// TIA Portal project "e009004v441" (V15.1)

(* hardware
DEVICE "Roll Forming"  TP1200 Comfort
   slot 0: "Roll Forming"  TP1200 Comfort  6AV2 124-0MC01-0AX0  15.1.0.0
   slot 1: "HMI_RT_1"  TP1200 Comfort  6AV2 124-0MC01-0AX0  15.1.0.0
   slot 5: "Roll Forming.IE_CP_1"  PROFINET Interface  15.0.1.0
      slot 1: "Interfaz PROFINET_1"  PROFINET Interface
         slot 1: "Port_1"  Port
         slot 2: "Port_2"  Port
   slot 7: "Roll Forming.MPI/DP_CP_1"  MPI/DP Interface  15.0.1.0
DEVICE "Dispositivo GSD_1"  GSD.Device
   slot 0: "Rack_0"  Rail
   slot 0: "Perfiladora"  6SL3 040-1MA00-0xxx  V4.3
DEVICE "PC-System_1"  SIMATIC PC station
   slot 0: "Estación PC SIMATIC"  Rail  SIMATIC PC-Station  V1.0
      slot 125: "Stationmanager"  Station_Manager  V6.0.4
   slot 1: "HMI_RT_2"  WinCC RT Advanced  6AV2 104-0xxxx-xxxx  15.1.0.0
      slot 33792: "Interfaz host"  Host interface
*)

(* ===== HMI "HMI_RT_1" =====

ScreenModuleEditorView "Bloc affichage_2" 800x600
   GraphicView "Affichage graphique" at 10,10 size 40x80; Picture "Graphique_9"
*)

(* ===== HMI "HMI_RT_1" =====
system functions are stored by id; their names below are inferred from use
connection "CPU 313C-2 DP": IF1 B, SIMATIC S7 300/400 MPI

HMI tags "Tabla de variables estándar"
   "DB_OP.COD2_ARRET" : DInt AT %DB50.DBD138, 1 s   // Encoder Formador 2 : Parar 1/10 mm
   "Desactivar_Falla59" : Bool AT %M87.2, 1 s
   "Desactivar_Falla78" : Bool AT %M89.5, 1 s
   "Desactivar_Falla47" : Bool AT %M85.6, 1 s
   "Desactivar_Falla84" : Bool AT %M90.3, 1 s
   "DB_OP.ACQ_DEFAUT" : Bool AT %DB50.DBX0.1, 1 s
   "Desactivar_Falla58" : Bool AT %M87.1, 1 s
   "Desactivar_Falla75" : Bool AT %M89.2, 1 s
   "35S2" : Bool AT %I12.1, 1 s   // Plegador 2 Fijación Abajo
   "28S3" : Bool AT %I5.2, 1 s   // Formador Herramienta 2 Matriz Off
   "Desactivar_Falla104" : Bool AT %M92.7, 1 s
   "Desactivar_Falla3" : Bool AT %M80.2, 1 s
   "Alarma_Cinta" : Bool AT %M96.4, 1 s
   "Desactivar_Falla68" : Bool AT %M88.3, 1 s
   "Desactivar_Falla38" : Bool AT %M84.5, 1 s
   "28S2" : Bool AT %I5.1, 1 s   // Formador Herramienta 2 Martillo On
   "DB_OP.COD1_VAL" : DInt AT %DB50.DBD100, 1 s   // Encoder Perfilador 1 : Valor 1/10 mm
   "31S3" : Bool AT %I8.2, 1 s   // Descargador Atrás
   "25S4" : Bool AT %I2.3, 1 s   // Pistón 1 Araña Contraído
   "Desactivar_Falla80" : Bool AT %M89.7, 1 s
   "Desactivar_Falla119" : Bool AT %M94.6, 1 s
   "Desactivar_Falla88" : Bool AT %M90.7, 1 s
   "HeladerasxMin" : Real AT %MD132, 1 s
   "Desactivar_Falla52" : Bool AT %M86.3, 1 s
   "Alarma_General" : Bool AT %M97.1, 1 s
   "DB_OP.DB_VAR" : Array [0..20] of Int AT %DB50.DBX8.0, 1 s   // Variables temporales
   "Desactivar_Falla11" : Bool AT %M81.2, 1 s
   "DB_OP.PI_COD_VAL" : DInt AT %DB50.DBD300, 1 s   // Encóder Pinza : Valor 1/10 mm
   "Desactivar_Falla116" : Bool AT %M94.3, 1 s
   "Desactivar_Falla102" : Bool AT %M92.5, 1 s
   "Hab_Medición" : Bool AT %M102.6, 1 s
   "35S3b" : Bool AT %I15.6, 1 s   // Plegador 2 posición Arriba (pata)
   "DB_OP.COD1_INIT" : DInt AT %DB50.DBD116, 1 s   // Encoder Perfilador 1 : Consigna Inicial 1/10 mm
   "Desactivar_Falla92" : Bool AT %M91.3, 1 s
   "28S8" : Bool AT %I5.7, 1 s   // Ajuste Formador Fin de Carrera Máx.
   "31S7b" : Bool AT %I15.5, 1 s   // Plegador 1 posición Arriba (pata)
   "DB_OP.COD2_CONS" : DInt AT %DB50.DBD134, 1 s   // Encoder Formador 2 : Consigna Posición 1/10 mm
   "DB_OP.DEF08" : Int AT %DB50.DBW94, 1 s   // IMAGE DEFAUT DBW 64
   "23S4" : Bool AT %I0.7, 1 s   // Presostato Freno Perfilador
   "Desactivar_Falla25" : Bool AT %M83.0, 1 s
   "Desactivar_Falla56" : Bool AT %M86.7, 1 s
   "DB_OP.DF_QM01" : Bool AT %DB50.DBX50.2, 1 s   // Térmico Intercambiador de Chapas
   "DB_OP.DEF06" : Int AT %DB50.DBW90, 1 s   // IMAGE DEFAUT DBW 60
   "DI8_CU_PL" : Bool AT %I62.7, 1 s   // Entrada Digital 8 CU Plegadores
   "DB_OP.DF_QM14" : Bool AT %DB50.DBX50.1, 1 s   // Térmico Calentador de Chapa
   "Desactivar_Falla39" : Bool AT %M84.6, 1 s
   "DB_OP.DEF01" : Int AT %DB50.DBW80, 1 s   // IMAGE DEFAUT DBW 50
   "32S5" : Bool AT %I9.4, 1 s   // Plegador 1 Extensión 2 Prensa Abajo
   "35S4_0" : Bool AT %I12.3, 1 s   // Plegador 2 Abajo
   "Desactivar_Falla112" : Bool AT %M93.7, 1 s
   "29S5" : Bool AT %I6.4, 1 s   // Pinza Cerrada
   "25S3" : Bool AT %I2.2, 1 s   // Fin de Carrera Araña Arriba
   "Desactivar_Falla93" : Bool AT %M91.4, 1 s
   "Desactivar_Falla111" : Bool AT %M93.6, 1 s
   "DB_OP.DF_QM06" : Bool AT %DB50.DBX51.2, 1 s   // Térmico Grupo Hidráulico Freno Perfilador
   "DB_OP.DF_VAR02" : Bool AT %DB50.DBX50.3, 1 s   // Defecto Vaiador Araña
   "30S3" : Bool AT %I7.2, 1 s   // Plegadora Tenaza arriba
   "Desactivar_Falla10" : Bool AT %M81.1, 1 s
   "DB_OP.PL2_COD_COEF" : Real AT %DB50.DBD262, 1 s   // Encoder Plegador 2 : Coeficiente Corrección
   "Desactivar_Falla6" : Bool AT %M80.5, 1 s
   "35S3" : Bool AT %I12.2, 1 s   // Plegador 2 Arriba
   "Desactivar_Falla103" : Bool AT %M92.6, 1 s
   "Alarma_Plegador" : Bool AT %M96.7, 1 s
   "DB_OP.PI_COD_DEC_PLI" : DInt AT %DB50.DBD322, 1 s   // Encóder Pinza : DECALAGE OUTIL PLIEUSE 1/10 mm
   "Desactivar_Falla36" : Bool AT %M84.3, 1 s
   "DB_OP.DF_LIM_PL1" : Bool AT %DB50.DBX51.7, 1 s   // Defecto Límite Plegador 1
   "Desactivar_Falla16" : Bool AT %M81.7, 1 s
   "26S4" : Bool AT %I3.3, 1 s   // Bajar Velocidad Transporte de Araña para Tomar Chapa
   "35S7" : Bool AT %I12.6, 1 s   // Plegador 2 Extensión 1 Prensa Abajo
   "27S4" : Bool AT %I4.3, 1 s   // Chapa en salida Perfilador
   "DB_OP.P_DEFAUT" : Bool AT %DB50.DBX0.0, 1 s
   "Desactivar_Falla71" : Bool AT %M88.6, 1 s
   "Desactivar_Falla48" : Bool AT %M85.7, 1 s
   "Desactivar_Falla125" : Bool AT %M95.4, 1 s
   "26S1" : Bool AT %I3.0, 1 s   // Tulipas no apoyadas en Chapa
   "DB_OP.COD1_CMD" : Bool AT %DB50.DBX128.0, 1 s   // Encoder Perfilador 1 : Inicio
   "30S7" : Bool AT %I7.6, 1 s   // Plegador 1 Cepillos Arriba
   "Desactivar_Falla83" : Bool AT %M90.2, 1 s
   "Alarma_Formador" : Bool AT %M96.5, 1 s
   "DB_OP.DEF05" : Int AT %DB50.DBW88, 1 s   // IMAGE DEFAUT DBW 58
   "Desactivar_Falla100" : Bool AT %M92.3, 1 s
   "21S6" : Bool AT %I124.7, 1 s   // Alineador Eje X Plegador 1 OFF
   "47K4" : Bool AT %Q8.3, 1 s   // Plegador 2 Bajar
   "Tiempo_Heladera_Prom" : Real AT %DB1.DBD40, 1 s
   "Desactivar_Falla107" : Bool AT %M93.2, 1 s
   "Desactivar_Falla114" : Bool AT %M94.1, 1 s
   "Desactivar_Falla21" : Bool AT %M82.4, 1 s
   "Desactivar_Falla31" : Bool AT %M83.6, 1 s
   "36S5" : Bool AT %I13.6, 1 s   // Plegador 2 Cepillos Arriba
   "29S4" : Bool AT %I6.3, 1 s   // Pinza Abierta
   "Desactivar_Falla97" : Bool AT %M92.0, 1 s
   "Desactivar_Falla14" : Bool AT %M81.5, 1 s
   "Desactivar_Falla82" : Bool AT %M90.1, 1 s
   "DB_OP.DF_LIM_PL2" : Bool AT %DB50.DBX52.0, 1 s   // Defecto Límite Plegador 2
   "Desactivar_Falla110" : Bool AT %M93.5, 1 s
   "35S2_0" : Bool AT %I12.1, 1 s   // Plegador 2 Fijación Abajo
   "Desactivar_Falla109" : Bool AT %M93.4, 1 s
   "Desactivar_Falla95" : Bool AT %M91.6, 1 s
   "36S6" : Bool AT %I13.7, 1 s   // Plegador 2 Cepillos Abajo
   "Desactivar_Falla76" : Bool AT %M89.3, 1 s
   "Selec_Pleg" : Int, internal
   "31S8" : Bool AT %I8.7, 1 s   // Plegador 1 Abajo
   "Alarma_Rolos" : Bool AT %M96.2, 1 s
   "27S6" : Bool AT %I4.5, 1 s   // Formador Herramienta 1 Martillo On
   "30S2" : Bool AT %I7.1, 1 s   // Plegadora Tenaza atrás
   "30S1" : Bool AT %I7.0, 1 s   // Plegadora Tenaza adelante
   "25S5" : Bool AT %I2.4, 1 s   // Fin de Carrera Araña Abajo
   "Desactivar_Falla29" : Bool AT %M83.4, 1 s
   "Desactivar_Falla13" : Bool AT %M81.4, 1 s
   "Desactivar_Falla23" : Bool AT %M82.6, 1 s
   "Alarma_Descargador" : Bool AT %M97.0, 1 s
   "DB_OP.PL1_COD_OFFSET" : DInt AT %DB50.DBD208, 1 s   // Encoder Plegador 1 : Consigna Inicial 1/10 mm
   "30S8" : Bool AT %I7.7, 1 s   // Plegador 1 Cepillos Abajo
   "DB_OP.PL2_COD_OFFSET" : DInt AT %DB50.DBD258, 1 s   // Encoder Plegador 2 : Consigna Inicial 1/10 mm
   "DB_OP.PI_COD_DEC_FORM" : DInt AT %DB50.DBD318, 1 s   // Encóder Pinza : DECALAGE OUTIL FORMAGE 1/10 mm
   "Alarma_Araña" : Bool AT %M96.1, 1 s
   "oHomming" : Bool AT %Q9.2, 1 s   // Lámpara Homming realizado
   "26S7" : Bool AT %I3.6, 1 s   // Presencia de Almacén 2 en Puesto de Trabajo
   "Simu Suelta Chapa" : Bool AT %M65.1, 1 s
   "Desactivar_Falla108" : Bool AT %M93.3, 1 s
   "DB_OP.COD2_COEF" : Real AT %DB50.DBD150, 1 s   // Encoder Formador 2 : Coeficiente Corrección
   "Ver_Tendencia" : Bool, internal
   "Desactivar_Falla46" : Bool AT %M85.5, 1 s
   "Desactivar_Falla40" : Bool AT %M84.7, 1 s
   "Simu Toma Chapa" : Bool AT %M65.0, 1 s
   "32S6" : Bool AT %I9.5, 1 s   // Plegador 1 Extensión 2 Prensa Arriba
   "Desactivar_Falla69" : Bool AT %M88.4, 1 s
   "35S3_0" : Bool AT %I12.2, 1 s   // Plegador 2 Arriba
   "35S5" : Bool AT %I12.4, 1 s   // Plegador 2 Prensa Abajo
   "Desactivar_Falla35" : Bool AT %M84.2, 1 s
   "26S3" : Bool AT %I3.2, 1 s   // Araña en Posición de Descarga
   "23S6" : Bool AT %I0.6, 1 s   // Alineador Eje Y Plegador 1 OFF
   "DB_OP.M2_P_CPT" : Int AT %DB50.DBW376, 1 s   // Almacén 2 Preselección contador de piezas
   "30S5" : Bool AT %I7.4, 1 s   // Plegadora Tenaza abierta
   "31S7" : Bool AT %I8.6, 1 s   // Plegador 1 Arriba
   "28S6" : Bool AT %I5.5, 1 s   // Matriz Formadora Bloqueo Herramienta Off
   "DB_OP.PL2_COD_CONS" : DInt AT %DB50.DBD254, 1 s   // Encoder Plegador 2 : Consigna Posición 1/10 mm
   "Desactivar_Falla62" : Bool AT %M87.5, 1 s
   "DB_OP.COD2_VAL" : DInt AT %DB50.DBD130, 1 s   // Encoder Formador 2 : Valor 1/10 mm
   "ProD" : DInt AT %MD200, 1 s
   "Tiempo_Heladera" : Real AT %MD136, 1 s
   "DB_OP.COD1_COEF" : Real AT %DB50.DBD120, 1 s   // Encoder Perfilador 1 : Coeficiente Corrección
   "23S5" : Bool AT %I0.5, 1 s   // Alineador Eje Y Plegador 1 ON
   "Desactivar_Falla26" : Bool AT %M83.1, 1 s
   "Desactivar_Falla79" : Bool AT %M89.6, 1 s
   "Desactivar_Falla63" : Bool AT %M87.6, 1 s
   "DB_OP.DEF02" : Int AT %DB50.DBW82, 1 s   // IMAGE DEFAUT DBW 52
   "Desactivar_Falla101" : Bool AT %M92.4, 1 s
   "Desactivar_Falla4" : Bool AT %M80.3, 1 s
   "Desactivar_Falla106" : Bool AT %M93.1, 1 s
   "25S8" : Bool AT %I2.7, 1 s   // Pistón 2 Araña Contraído
   "27S5" : Bool AT %I4.4, 1 s   // Formador Herramienta 1 Martillo Off
   "35S1" : Bool AT %I12.0, 1 s   // Plegador 2 Fijación Arriba
   "Desactivar_Falla61" : Bool AT %M87.4, 1 s
   "35S4" : Bool AT %I12.3, 1 s   // Plegador 2 Abajo
   "36S70" : Bool AT %I15.7, 1 s   // Barrera Atasco en Perfilador
   "Desactivar_Falla120" : Bool AT %M94.7, 1 s
   "32S4" : Bool AT %I9.3, 1 s   // Plegador 1 Extensión 1 Prensa Arriba
   "DB_OP.PL2_COD_VAL" : DInt AT %DB50.DBD250, 1 s   // Encoder Plegador 2 : Valor 1/10 mm
   "Desactivar_Falla64" : Bool AT %M87.7, 1 s
   "Desactivar_Falla43" : Bool AT %M85.2, 1 s
   "36S9" : Bool AT %I14.0, 1 s   // Plegador 1 Prensa en Posición Intermedia
   "32S2" : Bool AT %I9.1, 1 s   // Plegador 1 Prensa Arriba
   "DB_OP.RC2" : Int AT %DB50.DBW6, 1 s
   "25S7" : Bool AT %I2.6, 1 s   // Pistón 2 Araña Expandido
   "Desactivar_Falla17" : Bool AT %M82.0, 1 s
   "DB_OP.COD1_TARGET" : DInt AT %DB50.DBD112, 1 s   // Encoder Perfilador 1 : Ventana 1/10 mm
   "Desactivar_Falla54" : Bool AT %M86.5, 1 s
   "Desactivar_Falla9" : Bool AT %M81.0, 1 s
   "Desactivar_Falla53" : Bool AT %M86.4, 1 s
   "31S8_0" : Bool AT %I8.7, 1 s   // Plegador 1 Abajo
   "Desactivar_Falla67" : Bool AT %M88.2, 1 s
   "Alarma_Perfiladores" : Bool AT %M96.3, 1 s
   "21H1" : Bool AT %Q124.2, 1 s   // Lámpara En Ciclo
   "DB_OP.M2_V_CPT" : Int AT %DB50.DBW378, 1 s   // Almacén 2 contador de piezas
   "35S6" : Bool AT %I12.5, 1 s   // Plegador 2 Prensa Arriba
   "Desactivar_Falla7" : Bool AT %M80.6, 1 s
   "Desactivar_Falla121" : Bool AT %M95.0, 1 s
   "Desactivar_Falla27" : Bool AT %M83.2, 1 s
   "31S2" : Bool AT %I8.1, 1 s   // Descargador Adelante
   "Desactivar_Falla99" : Bool AT %M92.2, 1 s
   "Desactivar_Falla30" : Bool AT %M83.5, 1 s
   "45K7" : Bool AT %Q6.6, 1 s   // Subir Prensa Plegador 1
   "Desactivar_Falla86" : Bool AT %M90.5, 1 s
   "Desactivar_Falla74" : Bool AT %M89.1, 1 s
   "Desactivar_Falla15" : Bool AT %M81.6, 1 s
   "Desactivar_Falla98" : Bool AT %M92.1, 1 s
   "AjusteProF_Cinta" : Bool, internal
   "DB_OP.OP_SELMANU1" : Bool AT %DB50.DBX0.2, 1 s
   "Desactivar_Falla77" : Bool AT %M89.4, 1 s
   "30S6" : Bool AT %I7.5, 1 s   // Plegadora Tenaza cerrada
   "Desactivar_Falla94" : Bool AT %M91.5, 1 s
   "Reset_ProD" : Bool AT %M103.1, 1 s
   "Desactivar_Falla33" : Bool AT %M84.0, 1 s
   "DB_OP.COD1_CONS" : DInt AT %DB50.DBD104, 1 s   // Encoder Perfilador 1 : Consigna Posición 1/10 mm
   "Desactivar_Falla117" : Bool AT %M94.4, 1 s
   "32S3" : Bool AT %I9.2, 1 s   // Plegador 1 Extensión 1 Prensa Abajo
   "DB_OP.PL2_COD_VIT" : Int AT %DB50.DBW266, 1 s   // Encoder Plegador 2 : Velocidad Automática %
   "32S1" : Bool AT %I9.0, 1 s   // Plegador 1 Prensa Abajo
   "DB_OP.DF_QM13_2" : Bool AT %DB50.DBX50.0, 1 s   // Térmico Refrigeración Grupo Hidráulico
   "21S5" : Bool AT %I124.6, 1 s   // Alineador Eje X Plegador 1 ON
   "DB_OP.COD2_TARGET" : DInt AT %DB50.DBD142, 1 s   // Encoder Formador 2 : Ventana 1/10 mm
   "Desactivar_Falla65" : Bool AT %M88.0, 1 s
   "Desactivar_Falla70" : Bool AT %M88.5, 1 s
   "31S4" : Bool AT %I8.3, 1 s   // Barrera Seguridad Descargador
   "DB_OP.PI_COD_VIT1" : Int AT %DB50.DBW316, 1 s   // Encóder Pinza : Velocidad Automática %
   "Desactivar_Falla60" : Bool AT %M87.3, 1 s
   "28S4" : Bool AT %I5.3, 1 s   // Formador Herramienta 2 Matriz On
   "KM04_GV" : Bool AT %Q125.4, 1 s   // Velocidad Rápida Perfilador
   "Desactivar_Falla123" : Bool AT %M95.2, 1 s
   "Desactivar_Falla2" : Bool AT %M80.1, 1 s
   "DB_OP.COD2_CMD" : Bool AT %DB50.DBX158.0, 1 s   // Encoder Formador 2 : Inicio
   "DB_OP.M1_V_CPT" : Int AT %DB50.DBW374, 1 s   // Almacén 1 contador de piezas
   "Desactivar_Falla20" : Bool AT %M82.3, 1 s
   "Desactivar_Falla81" : Bool AT %M90.0, 1 s
   "Desactivar_Falla87" : Bool AT %M90.6, 1 s
   "31S5" : Bool AT %I8.4, 1 s   // Plegador 1 Fijación Arriba
   "Desactivar_Falla57" : Bool AT %M87.0, 1 s
   "Desactivar_Falla44" : Bool AT %M85.3, 1 s
   "29S3" : Bool AT %I6.2, 1 s   // Presencia de Chapa en Formador
   "36S8" : Bool AT %I13.1, 1 s   // Plegador 2 Extensión 2 Prensa Arriba
   "Desactivar_Falla66" : Bool AT %M88.1, 1 s
   "DB_OP.COD1_ARRET" : DInt AT %DB50.DBD108, 1 s   // Encoder Perfilador 1 : Parar 1/10 mm
   "Desactivar_Falla73" : Bool AT %M89.0, 1 s
   "DB_OP.DEF04" : Int AT %DB50.DBW86, 1 s   // IMAGE DEFAUT DBW 56
   "DB_OP.PL1_COD_CONS" : DInt AT %DB50.DBD204, 1 s   // Encoder Plegador 1 : Consigna Posición 1/10 mm
   "DB_OP.DEF07" : Int AT %DB50.DBW92, 1 s   // IMAGE DEFAUT DBW 62
   "26S2" : Bool AT %I3.1, 1 s   // Araña en Posicion de Carga
   "Desactivar_Falla90" : Bool AT %M91.1, 1 s
   "22S1_08" : Bool AT %I125.3, 1 s   // Rueda Unidades :8
   "Desactivar_Falla18" : Bool AT %M82.1, 1 s
   "Desactivar_Falla22" : Bool AT %M82.5, 1 s
   "26S5" : Bool AT %I3.4, 1 s   // Bajar Velocidad Transporte de Araña para Soltar Chapa
   "Desactivar_Falla41" : Bool AT %M85.0, 1 s
   "DB_OP.PL1_COD_VAL" : DInt AT %DB50.DBD200, 1 s   // Encoder Plegador 1 : Valor 1/10 mm
   "CA_47K5" : Bool AT %M22.6, 1 s   // Plegador 2 V1 Accionar
   "25S6" : Bool AT %I2.5, 1 s   // Araña Abajo
   "Desactivar_Falla89" : Bool AT %M91.0, 1 s
   "Desactivar_Falla37" : Bool AT %M84.4, 1 s
   "Desactivar_Falla124" : Bool AT %M95.3, 1 s
   "29S2" : Bool AT %I6.1, 1 s   // Formador Bloqueo de avance Off
   "Desactivar_Falla32" : Bool AT %M83.7, 1 s
   "Desactivar_Falla24" : Bool AT %M82.7, 1 s
   "36S1" : Bool AT %I13.2, 1 s   // Alineador Eje X Plegador 2 ON
   "27S7" : Bool AT %I4.6, 1 s   // Formador Herramienta 1 Matriz Off
   "26S8" : Bool AT %I3.7, 1 s   // Presencia de Chapa en Transporte Rolos
   "DB_OP.PI_COD_CONS" : DInt AT %DB50.DBD304, 1 s   // Encóder Pinza : Consigna Posición 1/10 mm
   "Desactivar_Falla49" : Bool AT %M86.0, 1 s
   "MANU" : Bool AT %M10.2, 1 s   // Modo Manual
      on ChangeValue: SetTag("Selec_Pleg", 0)
   "Desactivar_Falla12" : Bool AT %M81.3, 1 s
   "Alarma_Almacenes" : Bool AT %M96.0, 1 s
   "35S8" : Bool AT %I12.7, 1 s   // Plegador 2 Extensión 1 Prensa Arriba
   "30S4" : Bool AT %I7.3, 1 s   // Plegadora Tenaza abajo
   "Desactivar_Falla51" : Bool AT %M86.2, 1 s
   "Desactivar_Falla122" : Bool AT %M95.1, 1 s
   "Desactivar_Falla113" : Bool AT %M94.0, 1 s
   "DB_OP.PI_COD_COEF" : Real AT %DB50.DBD312, 1 s   // Encóder Pinza : Coeficiente Corrección
   "28S7" : Bool AT %I5.6, 1 s   // Ajuste Formador Fin de Carrera Mín.
   "29S7" : Bool AT %I6.6, 1 s   // Ajuste Ancho Perfilador Fin de carrera Máx.
   "DI9_CU_PL" : Bool AT %I82.7, 1 s   // Entrada Digital 9 CU Plegadores
   "Desactivar_Falla96" : Bool AT %M91.7, 1 s
   "28S1" : Bool AT %I5.0, 1 s   // Formador Herramienta 2 Martillo Off
   "Desactivar_Falla45" : Bool AT %M85.4, 1 s
   "32S6_0" : Bool AT %I9.5, 1 s   // Plegador 1 Extensión 2 Prensa Arriba
   "Desactivar_Falla34" : Bool AT %M84.1, 1 s
   "Desactivar_Falla42" : Bool AT %M85.1, 1 s
   "26S6" : Bool AT %I3.5, 1 s   // Presencia de Almacén 2 en Puesto de Espera
   "Desactivar_Falla1" : Bool AT %M80.0, 1 s
   "Desactivar_Falla28" : Bool AT %M83.3, 1 s
   "29S1" : Bool AT %I6.0, 1 s   // Formador Bloqueo de avance On
   "DB_OP.PL1_COD_VIT" : Int AT %DB50.DBW216, 1 s   // Encoder Plegador 1 : Velocidad Automática %
   "DB_OP.RC1" : Int AT %DB50.DBW4, 1 s
   "DB_OP.OP_SELMANU2" : Bool AT %DB50.DBX0.3, 1 s
   "DB_OP.PL1_COD1_RES1[13]" : Int AT %DB50.DBW242, 1 s   // Variable temporal
   "DB_OP.MODE" : Int AT %DB50.DBW2, 1 s   // Modo de Marcha
   "36S12" : Bool AT %I14.3, 1 s   // Descargador en Posición Intermedia
   "36S7" : Bool AT %I13.0, 1 s   // Plegador 2 Extensión 2 Prensa Abajo
   "Desactivar_Falla8" : Bool AT %M80.7, 1 s
   "AjusteProF_Perfiladores" : Bool, internal
   "DB_OP.COD2_INIT" : DInt AT %DB50.DBD146, 1 s   // Encoder Formador 2 : Consigna Inicial 1/10 mm
   "Desactivar_Falla118" : Bool AT %M94.5, 1 s
   "DB_OP.PI_COD_OFFSET" : DInt AT %DB50.DBD308, 1 s   // Encóder Pinza : Consigna Inicial 1/10 mm
   "HeladerasxHora" : Real AT %MD128, 1 s
   "Desactivar_Falla19" : Bool AT %M82.2, 1 s
   "Desactivar_Falla115" : Bool AT %M94.2, 1 s
   "Desactivar_Falla105" : Bool AT %M93.0, 1 s
   "Desactivar_Falla50" : Bool AT %M86.1, 1 s
   "Desactivar_Falla5" : Bool AT %M80.4, 1 s
   "28S5" : Bool AT %I5.4, 1 s   // Formador Bloqueo Herramienta On
   "Alarma_Pinza" : Bool AT %M96.6, 1 s
   "DB_OP.DEF03" : Int AT %DB50.DBW84, 1 s   // IMAGE DEFAUT DBW 54
   "Desactivar_Falla55" : Bool AT %M86.6, 1 s
   "Desactivar_Falla72" : Bool AT %M88.7, 1 s
   "36S2" : Bool AT %I13.3, 1 s   // Alineador Eje X Plegador 2 OFF
   "27S8" : Bool AT %I4.7, 1 s   // Formador Herramienta 1 Matriz On
   "DB_OP.M1_P_CPT" : Int AT %DB50.DBW372, 1 s   // Almacén 1 Preselección contador de piezas
   "31S6" : Bool AT %I8.5, 1 s   // Plegador 1 Fijación Abajo
   "DB_OP.PL1_COD_COEF" : Real AT %DB50.DBD212, 1 s   // Encoder Plegador 1 : Coeficiente Corrección
   "Desactivar_Falla85" : Bool AT %M90.4, 1 s
   "25S2" : Bool AT %I2.1, 1 s   // Desaceleración Transporte Cinta
   "Desactivar_Falla91" : Bool AT %M91.2, 1 s
   "27S3" : Bool AT %I4.2, 1 s   // Chapa en entrada Perfilador
   "IntentoResetFallido" : Bool AT %M110.0, 1 s
   "PosiciónFormado1" : DInt AT %DB53.DBD0, 1 s
   "PosiciónFormado2" : DInt AT %DB53.DBD4, 1 s
   "PosiciónFormado3" : DInt AT %DB53.DBD8, 1 s
   "PosiciónFormado4" : DInt AT %DB53.DBD12, 1 s
   "PL1_Pos01" : Bool AT %DB50.DBX393.1, 1 s
   "PL1_Pos02" : Bool AT %DB50.DBX393.2, 1 s
   "PL1_Pos03" : Bool AT %DB50.DBX393.3, 1 s
   "PL1_Pos04" : Bool AT %DB50.DBX393.4, 1 s
   "PL2_Pos00" : Bool AT %DB50.DBX394.0, 1 s
   "PL2_Pos01" : Bool AT %DB50.DBX394.1, 1 s
   "PL2_Pos02" : Bool AT %DB50.DBX394.2, 1 s
   "PL2_Pos03" : Bool AT %DB50.DBX394.3, 1 s
   "PL2_Pos04" : Bool AT %DB50.DBX394.4, 1 s
   "Pinza_Pos00" : Bool AT %DB50.DBX392.0, 1 s
   "Pinza_Pos01" : Bool AT %DB50.DBX392.1, 1 s
   "Pinza_Pos02" : Bool AT %DB50.DBX392.2, 1 s
   "Pinza_Pos03" : Bool AT %DB50.DBX392.3, 1 s
   "Pinza_Pos04" : Bool AT %DB50.DBX392.4, 1 s
   "Pinza_Pos05" : Bool AT %DB50.DBX392.5, 1 s
   "Comando_Inicializar_Araña" : Bool AT %M112.4, 1 s
   "Araña_Inicializada" : Bool AT %M112.3, 1 s
   "HommingPL1" : Bool AT %I62.6, 1 s
   "HommignPL2" : Bool AT %I82.6, 1 s
   "36S17" : Bool AT %I14.1, 1 s
   "29S6" : Bool AT %I6.5, 1 s
   "Hab_Almacenes" : Bool AT %M112.2, 1 s
   "Enclavamiento" : Bool AT %M0.5, 1 s
   "Warnings" : Byte AT %MB110, 1 s
   "Warning Activo" : Bool AT %M111.0, 1 s
   "Medición_Perf" : Real AT %DB2.DBD0, 1 s
   "Mostrar_Ajuste_Perf_1" : Bool, internal
   "Mostrar_Ajuste_Perf_2" : Bool, internal
   "Mostrar_Ajuste_Perf_3" : Bool, internal
   "eProC_Tiempos" : Bool, internal
   "HxHoraInst" : Real AT %DB1.DBD48, 1 s
   "Tiempo_Heladera_2" : Real AT %DB1.DBD4, 1 s
   "Tiempo_Heladera_3" : Real AT %DB1.DBD8, 1 s
   "Tiempo_Heladera_4" : Real AT %DB1.DBD12, 1 s
   "Tiempo_Heladera_5" : Real AT %DB1.DBD16, 1 s
   "Tiempo_Heladera_6" : Real AT %DB1.DBD20, 1 s
   "Tiempo_PL_Hid" : Real AT %DB1.DBD56, 1 s
   "Tiempo_PL_Neum" : Real AT %DB1.DBD60, 1 s
   "Tiempo_PL_Servos" : Real AT %DB1.DBD52, 1 s
   "Tiempo_PL_Descarga" : Real AT %DB1.DBD64, 1 s
   "Tiempo_PL_Descarga(parcial)" : Real AT %DB1.DBD80, 1 s
   "Tiempo_PL_Hid(parcial)" : Real AT %DB1.DBD72, 1 s
   "Tiempo_PL_Neum(parcial)" : Real AT %DB1.DBD76, 1 s
   "Tiempo_PL_Servos(parcial)" : Real AT %DB1.DBD68, 1 s
   "Tiempo_Heladera_Parcial" : Real AT %MD120, 1 s
   "Tiempo_Heladera_1" : Real AT %DB1.DBD0, 1 s
   "Ref_Pleg" : Bool AT %M62.5, 1 s
   "HabilitarReglasBaluff" : Bool AT %DB20.DBX24.0, 1 s
   "31S1" : Bool AT %I8.0, 1 s   // Presencia Producto en Descargador
   "SolRef_PL1" : Bool AT %DB21.DBX0.2, 1 s
   "SolRef_PL2" : Bool AT %DB21.DBX0.3, 1 s
   "Homing_PL1" : Bool AT %DB21.DBX0.0, 1 s
   "Homing_PL2" : Bool AT %DB21.DBX0.1, 1 s
   "HabRefPleg" : Bool AT %I15.4, 1 s
   "Descargador-ID_Bobina_Alm1" : DInt, internal
   "Descargador-ID_Bobina_Alm2" : DInt, internal
   "Descargador-FechaCorte_Alm1" : DateTime, internal
   "Descargador-FechaCorte_Alm2" : DateTime, internal
   "Contador_def_Alm1" : Int, internal
   "Contador_def_Alm2" : Int, internal
   "Defecto_Alm1" : Int, internal
   "Defecto_Alm2" : Int, internal
   "Proveedor_Indexado_Alm1" : Int, internal
   "Proveedor_Indexado_Alm2" : Int, internal

HMI tags "PiezaRolos"
   "Rolos\Rolos.C" : Int AT %DB7.DBW4, 1 s
   "Rolos\Rolos.PresenciaPieza" : Bool AT %DB7.DBX46.0, 1 s
   "Rolos\Rolos.PL2_2" : Int AT %DB7.DBW22, 1 s
   "Rolos\Actualizar2" : Bool AT %M65.3, 1 s
   "Rolos\Rolos.F3" : Int AT %DB7.DBW12, 1 s
   "Rolos\Rolos.D" : Int AT %DB7.DBW6, 1 s
   "Rolos\Rolos.F2" : Int AT %DB7.DBW10, 1 s
   "Rolos\Rolos.PL2_1" : Int AT %DB7.DBW20, 1 s
   "Rolos\Rolos.PL1_2" : Int AT %DB7.DBW18, 1 s
   "Rolos\Rolos.A" : Int AT %DB7.DBW0, 1 s
   "Rolos\Actualizar" : Bool AT %M65.2, 1 s
   "Rolos\Rolos.F4" : Int AT %DB7.DBW14, 1 s
   "Rolos\Rolos.B" : Int AT %DB7.DBW2, 1 s
   "Rolos\Rolos.F1" : Int AT %DB7.DBW8, 1 s
   "Rolos\Rolos.PL1_1" : Int AT %DB7.DBW16, 1 s
   "Rolos\Rolos.Nombre" : String[20] AT %DB7.DBX24.0, 1 s

HMI tags "PiezaPinza"
   "Pinza\Pinza.F4" : Int AT %DB10.DBW14, 1 s
   "Pinza\Pinza.F2" : Int AT %DB10.DBW10, 1 s
   "Pinza\Pinza.PL2_1" : Int AT %DB10.DBW20, 1 s
   "Pinza\Pinza.PL2_2" : Int AT %DB10.DBW22, 1 s
   "Pinza\Pinza.B" : Int AT %DB10.DBW2, 1 s
   "Pinza\Pinza.PresenciaPieza" : Bool AT %DB10.DBX46.0, 1 s
   "Pinza\Pinza.PL1_2" : Int AT %DB10.DBW18, 1 s
   "Pinza\Pinza.F1" : Int AT %DB10.DBW8, 1 s
   "Pinza\Pinza.A" : Int AT %DB10.DBW0, 1 s
   "Pinza\Pinza.F3" : Int AT %DB10.DBW12, 1 s
   "Pinza\Pinza.C" : Int AT %DB10.DBW4, 1 s
   "Pinza\Pinza.PL1_1" : Int AT %DB10.DBW16, 1 s
   "Pinza\Pinza.D" : Int AT %DB10.DBW6, 1 s
   "Pinza\Pinza.Nombre" : String[20] AT %DB10.DBX24.0, 1 s

HMI tags "PiezaPlegadores"
   "Plegadora\Plegadora.F4" : Int AT %DB11.DBW14, 1 s
   "Plegadora\Plegadora.PresenciaPieza" : Bool AT %DB11.DBX46.0, 1 s
   "Plegadora\Plegadora.B" : Int AT %DB11.DBW2, 1 s
   "Plegadora\Plegadora.F1" : Int AT %DB11.DBW8, 1 s
   "Plegadora\Plegadora.A" : Int AT %DB11.DBW0, 1 s
   "Plegadora\Plegadora.C" : Int AT %DB11.DBW4, 1 s
   "Plegadora\Plegadora.F3" : Int AT %DB11.DBW12, 1 s
   "Plegadora\Plegadora.PL2_1" : Int AT %DB11.DBW20, 1 s
   "Plegadora\Plegadora.PL1_1" : Int AT %DB11.DBW16, 1 s
   "Plegadora\Plegadora.F2" : Int AT %DB11.DBW10, 1 s
   "Plegadora\Plegadora.PL1_2" : Int AT %DB11.DBW18, 1 s
   "Plegadora\Plegadora.D" : Int AT %DB11.DBW6, 1 s
   "Plegadora\Plegadora.PL2_2" : Int AT %DB11.DBW22, 1 s
   "Plegadora\Plegadora.Nombre" : String[20] AT %DB11.DBX24.0, 1 s

HMI tags "PiezaAraña"
   "Araña\Araña.PresenciaPieza" : Bool AT %DB6.DBX46.0, 1 s
   "Araña\Araña.F4" : Int AT %DB6.DBW14, 1 s
   "Araña\Araña.B" : Int AT %DB6.DBW2, 1 s
   "Araña\Araña.C" : Int AT %DB6.DBW4, 1 s
   "Araña\Araña.PL2_1" : Int AT %DB6.DBW20, 1 s
   "Araña\Araña.PL1_1" : Int AT %DB6.DBW16, 1 s
   "Araña\Araña.A" : Int AT %DB6.DBW0, 1 s
   "Araña\Actualizar2" : Bool AT %M65.1, 1 s
   "Araña\Araña.F2" : Int AT %DB6.DBW10, 1 s
   "Araña\Actualizar" : Bool AT %M65.0, 1 s
   "Araña\Araña.PL1_2" : Int AT %DB6.DBW18, 1 s
   "Araña\Araña.PL2_2" : Int AT %DB6.DBW22, 1 s
   "Araña\Araña.F1" : Int AT %DB6.DBW8, 1 s
   "Araña\Araña.F3" : Int AT %DB6.DBW12, 1 s
   "Araña\Araña.D" : Int AT %DB6.DBW6, 1 s
   "Araña\Araña.Nombre" : String[20] AT %DB6.DBX24.0, 1 s

HMI tags "PiezaReceta"
   "Receta\Recetas.A" : Int AT %DB3.DBW0, 1 s   // Mot Piece : Côte A
   "Receta\Recetas.PL2_1" : Int AT %DB3.DBW20, 1 s   // Plegador 2 Pliego 1
   "Receta\Recetas.F2" : Int AT %DB3.DBW10, 1 s   // Punto de Formado 2
   "Receta\Recetas.F1" : Int AT %DB3.DBW8, 1 s   // Punto de Formado 1
   "Receta\Recetas.PL2_2" : Int AT %DB3.DBW22, 1 s   // Plegador 2 Pliego 2
   "Receta\Recetas.x_M1" : Bool AT %M180.7, 1 s   // BP _tranfert reference sur magasin 1
   "Receta\Recetas.F4" : Int AT %DB3.DBW14, 1 s   // Punto de Formado 4
   "Receta\Recetas.D" : Int AT %DB3.DBW6, 1 s   // Mot Piece : Côte D
   "Receta\Recetas.F3" : Int AT %DB3.DBW12, 1 s   // Punto de Formado 3
   "Receta\VerHeladera" : Bool, internal
   "Receta\Recetas.x_M2" : Bool AT %M181.0, 1 s   // BP _tranfert reference sur magasin 2
   "Receta\Recetas.Nombre" : String[20] AT %DB3.DBX24.0, 1 s
   "Receta\Recetas.B" : Int AT %DB3.DBW2, 1 s   // Mot Piece : Côte B
   "Receta\Recetas.PL1_2" : Int AT %DB3.DBW18, 1 s   // Plegador 1 Pliego 2
   "Receta\Recetas.PL1_1" : Int AT %DB3.DBW16, 1 s   // Plegador 1 Pliego 1
   "Receta\Recetas.C" : Int AT %DB3.DBW4, 1 s   // Mot Piece : Côte C

HMI tags "Tag table_6"
   "Receta Almacén1\OFFSET.REC_MG1.OFFSET_F2" : Int AT %DB52.DBW32, 1 s   // Punto de Formado 2
   "Receta Almacén1\OFFSET.REC_MG1.OFFSET_F4" : Int AT %DB52.DBW36, 1 s   // Punto de Formado 4
   "Receta Almacén1\OFFSET.REC_MG1.OFFSET_PL1_1" : Int AT %DB52.DBW38, 1 s   // Plegador 1 Pliego 1
   "Receta Almacén1\OFFSET.REC_MG1.OFFSET_PL2_1" : Int AT %DB52.DBW42, 1 s   // Plegador 2 Pliego 1
   "Receta Almacén1\DB_OP.M1.MPP" : Bool AT %DB50.DBX400.0, 1 s   // Presencia de Pieza
   "Receta Almacén1\Recetas.REC_MG1.NOM" : String[8] AT %DB51.DBX130.0, 1 s
   "Receta Almacén1\DB_OP.M1T_XCPT" : Bool AT %DB50.DBX380.0, 1 s   // Almacén 1 Entrega Pieza
   "Receta Almacén1\VerHeladera" : Bool, internal
   "Receta Almacén1\Recetas.REC_MG1.A_0" : DInt AT %DB51.DBD148, 1 s   // Mot Piece : Côte B
   "Receta Almacén1\OFFSET.REC_MG1.OFFSET_PL1_2" : Int AT %DB52.DBW40, 1 s   // Plegador 1 Pliego 2
   "Receta Almacén1\Detalles" : Bool, internal
   "Receta Almacén1\Recetas.REC_MG1.A" : DInt AT %DB51.DBD144, 1 s   // Mot Piece : Côte A
   "Receta Almacén1\OFFSET.REC_MG1.OFFSET_F3" : Int AT %DB52.DBW34, 1 s   // Punto de Formado 3
   "Receta Almacén1\OFFSET.REC_MG1.OFFSET_PL2_2" : Int AT %DB52.DBW44, 1 s   // Plegador 2 Pliego 2
   "Receta Almacén1\OFFSET.REC_MG1.OFFSET_F1" : Int AT %DB52.DBW30, 1 s   // Punto de Formado 1
   "Receta Almacén1\26S7" : Bool AT %I3.6, 1 s   // Presencia de Almacén 2 en Puesto de Trabajo
   "Receta Almacén1\CA_KM01_1" : Bool AT %M18.4, 1 s   // Intercambiador Almacenes Avance (Alm1)
   "Receta Almacén1\Recetas.REC_MG1.D" : DInt AT %DB51.DBD156, 1 s   // Mot Piece : Côte D
   "Receta Almacén1\Recetas.REC_MG1.C" : DInt AT %DB51.DBD152, 1 s   // Mot Piece : Côte C
